// TIA Portal project "OP-TQ-01" (V13) (continued)
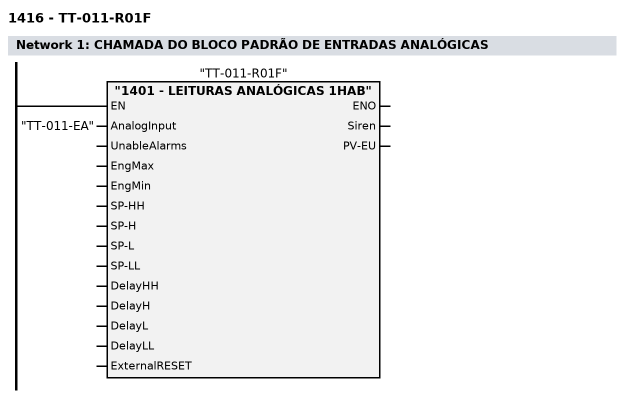
   RUNG wire#powerrail
      "TT-011-R01F"(AnalogInput := "TT-011-EA", UnableAlarms :=, EngMax :=, EngMin :=, "SP-HH" :=, "SP-H" :=, "SP-L" :=, "SP-LL" :=, DelayHH :=, DelayH :=, DelayL :=, DelayLL :=, ExternalRESET :=, Siren =>, "PV-EU" =>)
   END_RUNG
   // the same network as SCL:
   "TT-011-R01F"(AnalogInput := "TT-011-EA");   // "1401 - LEITURAS ANALÓGICAS 1HAB"
END_REGION
END_FUNCTION

// folder: PARAMETRIZADOS

FUNCTION_BLOCK "1110 - RESISTENCIAS"   // FB1110, LAD
{ S7_Optimized_Access := 'FALSE' }
VERSION : 0.1
   VAR_TEMP   // added for the SCL form of the ladder/FBD networks
      _w1 : Bool;
      _w2 : Bool;
   END_VAR
BEGIN

REGION Network 1: RESET FALHAS
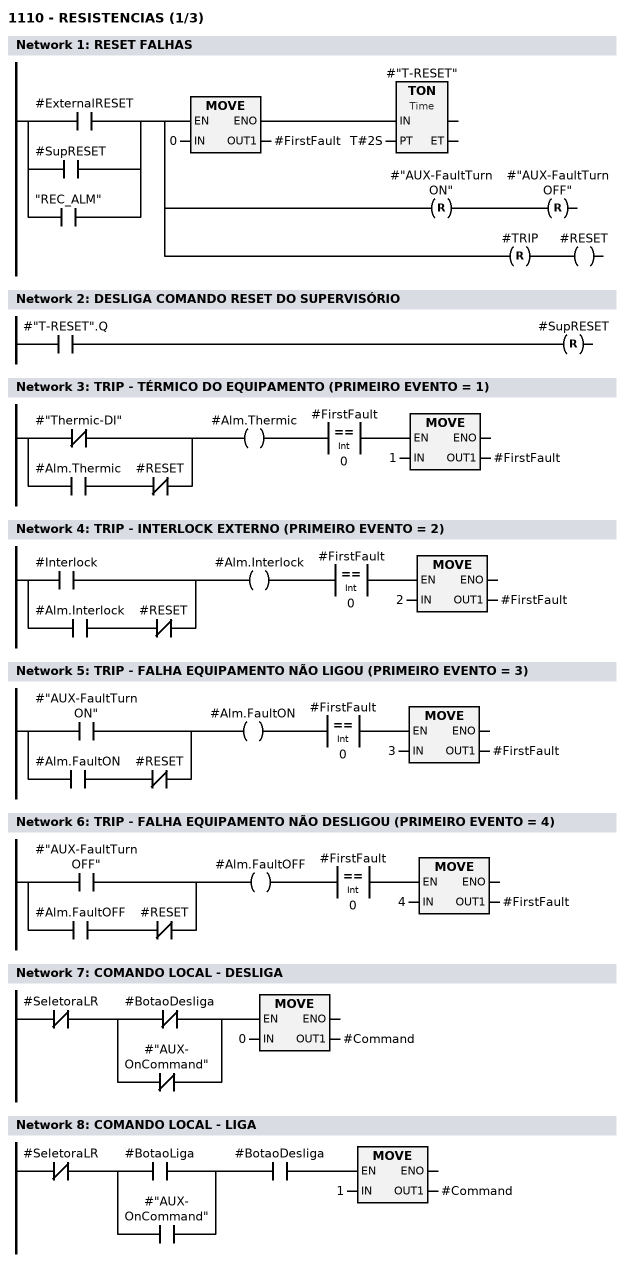
   // ENO of a box is taken as its EN; it also drops when the box reports an error
   #_w1 := #ExternalRESET OR #SupRESET OR "REC_ALM";
   IF #_w1 THEN #FirstFault := 0; END_IF;
   #"T-RESET".TON(IN := #_w1, PT := T#2S);
   IF #_w1 THEN
       #"AUX-FaultTurnON" := FALSE;
       #"AUX-FaultTurnOFF" := FALSE;
       #TRIP := FALSE;
   END_IF;
   #RESET := #_w1;
END_REGION

REGION Network 2: DESLIGA COMANDO RESET DO SUPERVISÓRIO
   RUNG wire#powerrail
      Contact( #"T-RESET".Q )
      R_Coil( #SupRESET )
   END_RUNG
   // the same network as SCL:
   IF #"T-RESET".Q THEN #SupRESET := FALSE; END_IF;
END_REGION

REGION Network 3: TRIP - TÉRMICO DO EQUIPAMENTO (PRIMEIRO EVENTO = 1)
   RUNG wire#powerrail
      I_Contact( #"Thermic-DI" )
      wire#w1
      Coil( #Alm.Thermic )
      { S7_Templates := "SrcType := Int" } EQ_Contact(in1 := #FirstFault, in2 := 0)
      { S7_GenerateENO := "TRUE" } Move(in := 1, out1 => #FirstFault)
   END_RUNG
   RUNG wire#powerrail
      Contact( #Alm.Thermic )
      I_Contact( #RESET )
   END_RUNG wire#w1
   // the same network as SCL:
   #Alm.Thermic := NOT #"Thermic-DI" OR (#Alm.Thermic AND NOT #RESET);
   IF #Alm.Thermic AND (#FirstFault = 0) THEN #FirstFault := 1; END_IF;
END_REGION

REGION Network 4: TRIP - INTERLOCK EXTERNO (PRIMEIRO EVENTO = 2)
   RUNG wire#powerrail
      Contact( #Interlock )
      wire#w1
      Coil( #Alm.Interlock )
      { S7_Templates := "SrcType := Int" } EQ_Contact(in1 := #FirstFault, in2 := 0)
      { S7_GenerateENO := "TRUE" } Move(in := 2, out1 => #FirstFault)
   END_RUNG
   RUNG wire#powerrail
      Contact( #Alm.Interlock )
      I_Contact( #RESET )
   END_RUNG wire#w1
   // the same network as SCL:
   #Alm.Interlock := #Interlock OR (#Alm.Interlock AND NOT #RESET);
   IF #Alm.Interlock AND (#FirstFault = 0) THEN #FirstFault := 2; END_IF;
END_REGION

REGION Network 5: TRIP - FALHA EQUIPAMENTO NÃO LIGOU (PRIMEIRO EVENTO = 3)
   RUNG wire#powerrail
      Contact( #"AUX-FaultTurnON" )
      wire#w1
      Coil( #Alm.FaultON )
      { S7_Templates := "SrcType := Int" } EQ_Contact(in1 := #FirstFault, in2 := 0)
      { S7_GenerateENO := "TRUE" } Move(in := 3, out1 => #FirstFault)
   END_RUNG
   RUNG wire#powerrail
      Contact( #Alm.FaultON )
      I_Contact( #RESET )
   END_RUNG wire#w1
   // the same network as SCL:
   #Alm.FaultON := #"AUX-FaultTurnON" OR (#Alm.FaultON AND NOT #RESET);
   IF #Alm.FaultON AND (#FirstFault = 0) THEN #FirstFault := 3; END_IF;
END_REGION

REGION Network 6: TRIP - FALHA EQUIPAMENTO NÃO DESLIGOU (PRIMEIRO EVENTO = 4)
   RUNG wire#powerrail
      Contact( #"AUX-FaultTurnOFF" )
      wire#w1
      Coil( #Alm.FaultOFF )
      { S7_Templates := "SrcType := Int" } EQ_Contact(in1 := #FirstFault, in2 := 0)
      { S7_GenerateENO := "TRUE" } Move(in := 4, out1 => #FirstFault)
   END_RUNG
   RUNG wire#powerrail
      Contact( #Alm.FaultOFF )
      I_Contact( #RESET )
   END_RUNG wire#w1
   // the same network as SCL:
   #Alm.FaultOFF := #"AUX-FaultTurnOFF" OR (#Alm.FaultOFF AND NOT #RESET);
   IF #Alm.FaultOFF AND (#FirstFault = 0) THEN #FirstFault := 4; END_IF;
END_REGION

REGION Network 7: COMANDO LOCAL - DESLIGA
   RUNG wire#powerrail
      I_Contact( #SeletoraLR )
      wire#w1
      I_Contact( #BotaoDesliga )
      wire#w2
      { S7_GenerateENO := "TRUE" } Move(in := 0, out1 => #Command)
   END_RUNG
   RUNG wire#w1
      I_Contact( #"AUX-OnCommand" )
   END_RUNG wire#w2
   // the same network as SCL:
   IF NOT #SeletoraLR AND (NOT #BotaoDesliga OR NOT #"AUX-OnCommand") THEN #Command := 0; END_IF;
END_REGION

REGION Network 8: COMANDO LOCAL - LIGA
   RUNG wire#powerrail
      I_Contact( #SeletoraLR )
      wire#w1
      Contact( #BotaoLiga )
      wire#w2
      Contact( #BotaoDesliga )
      { S7_GenerateENO := "TRUE" } Move(in := 1, out1 => #Command)
   END_RUNG
   RUNG wire#w1
      Contact( #"AUX-OnCommand" )
   END_RUNG wire#w2
   // the same network as SCL:
   IF NOT #SeletoraLR AND (#BotaoLiga OR #"AUX-OnCommand") AND #BotaoDesliga THEN #Command := 1; END_IF;
END_REGION

REGION Network 9: COMANDO LIGA EQUIPAMENTO
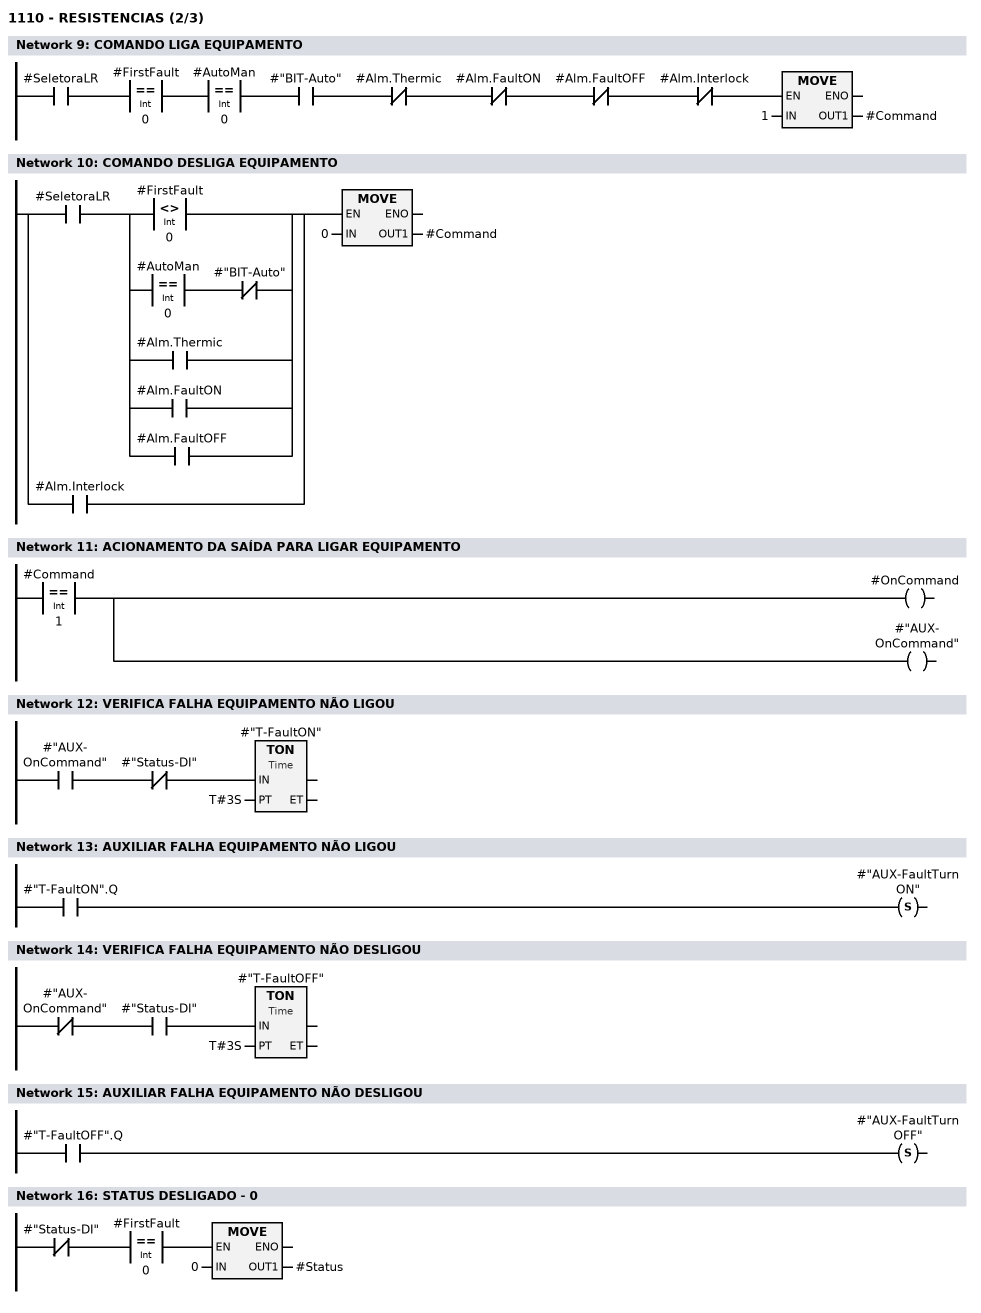
   RUNG wire#powerrail
      Contact( #SeletoraLR )
      { S7_Templates := "SrcType := Int" } EQ_Contact(in1 := #FirstFault, in2 := 0)
      { S7_Templates := "SrcType := Int" } EQ_Contact(in1 := #AutoMan, in2 := 0)
      Contact( #"BIT-Auto" )
      I_Contact( #Alm.Thermic )
      I_Contact( #Alm.FaultON )
      I_Contact( #Alm.FaultOFF )
      I_Contact( #Alm.Interlock )
      { S7_GenerateENO := "TRUE" } Move(in := 1, out1 => #Command)
   END_RUNG
   // the same network as SCL:
   IF #SeletoraLR AND (#FirstFault = 0) AND (#AutoMan = 0) AND #"BIT-Auto" AND NOT #Alm.Thermic AND NOT #Alm.FaultON AND NOT #Alm.FaultOFF AND NOT #Alm.Interlock THEN
       #Command := 1;
   END_IF;
END_REGION

REGION Network 10: COMANDO DESLIGA EQUIPAMENTO
   RUNG wire#powerrail
      Contact( #SeletoraLR )
      wire#w1
      { S7_Templates := "SrcType := Int" } NE_Contact(in1 := #FirstFault, in2 := 0)
      wire#w2
      { S7_GenerateENO := "TRUE" } Move(in := 0, out1 => #Command)
   END_RUNG
   RUNG wire#w1
      { S7_Templates := "SrcType := Int" } EQ_Contact(in1 := #AutoMan, in2 := 0)
      I_Contact( #"BIT-Auto" )
   END_RUNG wire#w2
   RUNG wire#w1
      Contact( #Alm.Thermic )
   END_RUNG wire#w2
   RUNG wire#w1
      Contact( #Alm.FaultON )
   END_RUNG wire#w2
   RUNG wire#w1
      Contact( #Alm.FaultOFF )
   END_RUNG wire#w2
   RUNG wire#powerrail
      Contact( #Alm.Interlock )
   END_RUNG wire#w2
   // the same network as SCL:
   IF (#SeletoraLR AND ((#FirstFault <> 0) OR ((#AutoMan = 0) AND NOT #"BIT-Auto") OR #Alm.Thermic OR #Alm.FaultON OR #Alm.FaultOFF)) OR #Alm.Interlock THEN
       #Command := 0;
   END_IF;
END_REGION

REGION Network 11: ACIONAMENTO DA SAÍDA PARA LIGAR EQUIPAMENTO
   RUNG wire#powerrail
      { S7_Templates := "SrcType := Int" } EQ_Contact(in1 := #Command, in2 := 1)
      wire#w1
      Coil( #OnCommand )
   END_RUNG
   RUNG wire#w1
      Coil( #"AUX-OnCommand" )
   END_RUNG
   // the same network as SCL:
   #OnCommand := #Command = 1;
   #"AUX-OnCommand" := #OnCommand;
END_REGION

REGION Network 12: VERIFICA FALHA EQUIPAMENTO NÃO LIGOU
   #"T-FaultON".TON(IN := #"AUX-OnCommand" AND NOT #"Status-DI", PT := T#3S);
END_REGION

REGION Network 13: AUXILIAR FALHA EQUIPAMENTO NÃO LIGOU
   RUNG wire#powerrail
      Contact( #"T-FaultON".Q )
      S_Coil( #"AUX-FaultTurnON" )
   END_RUNG
   // the same network as SCL:
   IF #"T-FaultON".Q THEN #"AUX-FaultTurnON" := TRUE; END_IF;
END_REGION

REGION Network 14: VERIFICA FALHA EQUIPAMENTO NÃO DESLIGOU
   #"T-FaultOFF".TON(IN := NOT #"AUX-OnCommand" AND #"Status-DI", PT := T#3S);
END_REGION

REGION Network 15: AUXILIAR FALHA EQUIPAMENTO NÃO DESLIGOU
   RUNG wire#powerrail
      Contact( #"T-FaultOFF".Q )
      S_Coil( #"AUX-FaultTurnOFF" )
   END_RUNG
   // the same network as SCL:
   IF #"T-FaultOFF".Q THEN #"AUX-FaultTurnOFF" := TRUE; END_IF;
END_REGION

REGION Network 16: STATUS DESLIGADO - 0
   RUNG wire#powerrail
      I_Contact( #"Status-DI" )
      { S7_Templates := "SrcType := Int" } EQ_Contact(in1 := #FirstFault, in2 := 0)
      { S7_GenerateENO := "TRUE" } Move(in := 0, out1 => #Status)
   END_RUNG
   // the same network as SCL:
   IF NOT #"Status-DI" AND (#FirstFault = 0) THEN #Status := 0; END_IF;
END_REGION

REGION Network 17: STATUS LIGADO - 1
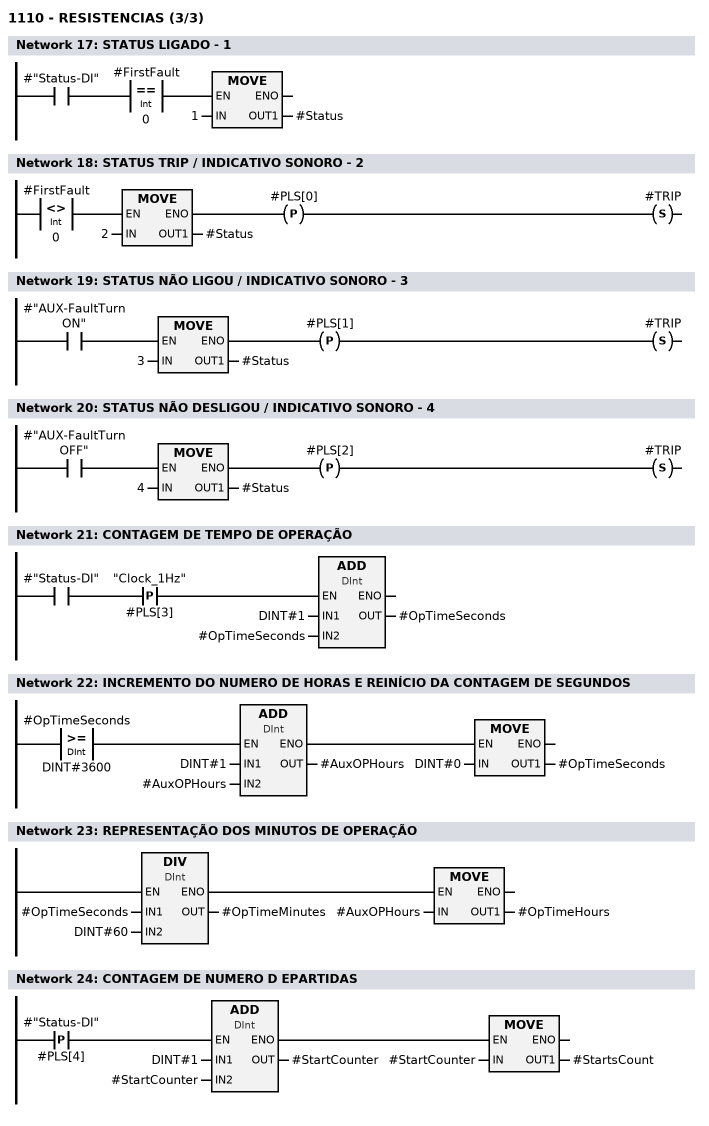
   RUNG wire#powerrail
      Contact( #"Status-DI" )
      { S7_Templates := "SrcType := Int" } EQ_Contact(in1 := #FirstFault, in2 := 0)
      { S7_GenerateENO := "TRUE" } Move(in := 1, out1 => #Status)
   END_RUNG
   // the same network as SCL:
   IF #"Status-DI" AND (#FirstFault = 0) THEN #Status := 1; END_IF;
END_REGION

REGION Network 18: STATUS TRIP / INDICATIVO SONORO - 2
   RUNG wire#powerrail
      { S7_Templates := "SrcType := Int" } NE_Contact(in1 := #FirstFault, in2 := 0)
      { S7_GenerateENO := "TRUE" } Move(in := 2, out1 => #Status)
      P_Trig( #PLS[0] )
      S_Coil( #TRIP )
   END_RUNG
   // the same network as SCL:
   // ENO of a box is taken as its EN; it also drops when the box reports an error
   #_w1 := #FirstFault <> 0;
   IF #_w1 THEN #Status := 2; END_IF;
   #_w2 := #_w1 AND NOT #PLS[0];   // rising edge
   #PLS[0] := #_w1;
   IF #_w2 THEN #TRIP := TRUE; END_IF;
END_REGION

REGION Network 19: STATUS NÃO LIGOU / INDICATIVO SONORO - 3
   RUNG wire#powerrail
      Contact( #"AUX-FaultTurnON" )
      { S7_GenerateENO := "TRUE" } Move(in := 3, out1 => #Status)
      P_Trig( #PLS[1] )
      S_Coil( #TRIP )
   END_RUNG
   // the same network as SCL:
   // ENO of a box is taken as its EN; it also drops when the box reports an error
   IF #"AUX-FaultTurnON" THEN #Status := 3; END_IF;
   #_w1 := #"AUX-FaultTurnON" AND NOT #PLS[1];   // rising edge
   #PLS[1] := #"AUX-FaultTurnON";
   IF #_w1 THEN #TRIP := TRUE; END_IF;
END_REGION

REGION Network 20: STATUS NÃO DESLIGOU / INDICATIVO SONORO - 4
   RUNG wire#powerrail
      Contact( #"AUX-FaultTurnOFF" )
      { S7_GenerateENO := "TRUE" } Move(in := 4, out1 => #Status)
      P_Trig( #PLS[2] )
      S_Coil( #TRIP )
   END_RUNG
   // the same network as SCL:
   // ENO of a box is taken as its EN; it also drops when the box reports an error
   IF #"AUX-FaultTurnOFF" THEN #Status := 4; END_IF;
   #_w1 := #"AUX-FaultTurnOFF" AND NOT #PLS[2];   // rising edge
   #PLS[2] := #"AUX-FaultTurnOFF";
   IF #_w1 THEN #TRIP := TRUE; END_IF;
END_REGION

REGION Network 21: CONTAGEM DE TEMPO DE OPERAÇÃO
   RUNG wire#powerrail
      Contact( #"Status-DI" )
      P_Contact(operand := "Clock_1Hz", bit := #PLS[3])
      { S7_Templates := "SrcType := DInt"; S7_GenerateENO := "TRUE" } Add(in1 := DINT#1, in2 := #OpTimeSeconds, out => #OpTimeSeconds)
   END_RUNG
   // the same network as SCL:
   #_w1 := #"Status-DI" AND "Clock_1Hz" AND NOT #PLS[3];   // rising edge of "Clock_1Hz"
   #PLS[3] := "Clock_1Hz";
   IF #_w1 THEN #OpTimeSeconds := DINT#1 + #OpTimeSeconds; END_IF;
END_REGION

REGION Network 22: INCREMENTO DO NUMERO DE HORAS E REINÍCIO DA CONTAGEM DE SEGUNDOS
   RUNG wire#powerrail
      { S7_Templates := "SrcType := DInt" } GE_Contact(in1 := #OpTimeSeconds, in2 := DINT#3600)
      { S7_Templates := "SrcType := DInt"; S7_GenerateENO := "TRUE" } Add(in1 := DINT#1, in2 := #AuxOPHours, out => #AuxOPHours)
      { S7_GenerateENO := "TRUE" } Move(in := DINT#0, out1 => #OpTimeSeconds)
   END_RUNG
   // the same network as SCL:
   // ENO of a box is taken as its EN; it also drops when the box reports an error
   IF #OpTimeSeconds >= DINT#3600 THEN
       #AuxOPHours := DINT#1 + #AuxOPHours;
       #OpTimeSeconds := DINT#0;
   END_IF;
END_REGION

REGION Network 23: REPRESENTAÇÃO DOS MINUTOS DE OPERAÇÃO
   RUNG wire#powerrail
      { S7_Templates := "SrcType := DInt"; S7_GenerateENO := "TRUE" } Div(in1 := #OpTimeSeconds, in2 := DINT#60, out => #OpTimeMinutes)
      { S7_GenerateENO := "TRUE" } Move(in := #AuxOPHours, out1 => #OpTimeHours)
   END_RUNG
   // the same network as SCL:
   // ENO of a box is taken as its EN; it also drops when the box reports an error
   #OpTimeMinutes := #OpTimeSeconds / DINT#60;
   #OpTimeHours := #AuxOPHours;
END_REGION

REGION Network 24: CONTAGEM DE NUMERO D EPARTIDAS
   RUNG wire#powerrail
      P_Contact(operand := #"Status-DI", bit := #PLS[4])
      { S7_Templates := "SrcType := DInt"; S7_GenerateENO := "TRUE" } Add(in1 := DINT#1, in2 := #StartCounter, out => #StartCounter)
      { S7_GenerateENO := "TRUE" } Move(in := #StartCounter, out1 => #StartsCount)
   END_RUNG
   // the same network as SCL:
   // ENO of a box is taken as its EN; it also drops when the box reports an error
   #_w1 := #"Status-DI" AND NOT #PLS[4];   // rising edge of #"Status-DI"
   #PLS[4] := #"Status-DI";
   IF #_w1 THEN
       #StartCounter := DINT#1 + #StartCounter;
       #StartsCount := #StartCounter;
   END_IF;
END_REGION
END_FUNCTION_BLOCK

FUNCTION_BLOCK "1401 - LEITURAS ANALÓGICAS 1HAB"   // FB1401, LAD
TITLE = LEITURA E VERIFICAÇÃO DE ALARMES ANALÓGICOS
{ S7_Optimized_Access := 'FALSE' }
VERSION : 0.1
   VAR_TEMP   // added for the SCL form of the ladder/FBD networks
      _w1 : Bool;
      _w2 : Bool;
      _w3 : Bool;
      _w4 : Bool;
   END_VAR
BEGIN

REGION Network 1: RESET FALHAS
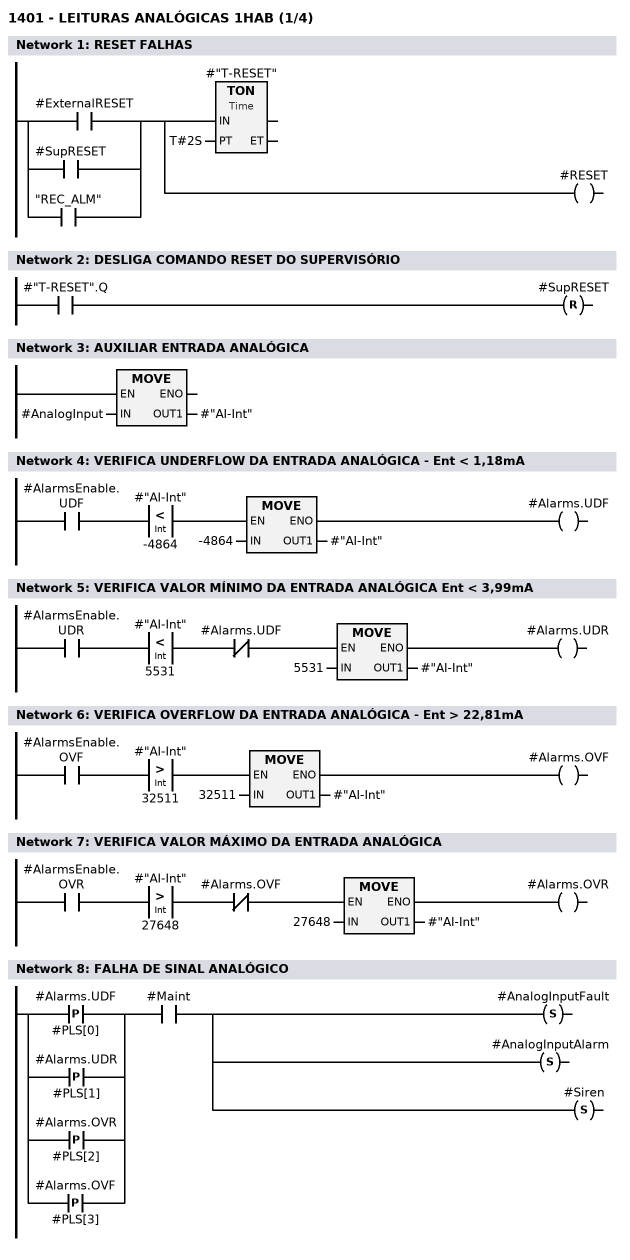
   #_w1 := #ExternalRESET OR #SupRESET OR "REC_ALM";
   #"T-RESET".TON(IN := #_w1, PT := T#2S);
   #RESET := #_w1;
END_REGION

REGION Network 2: DESLIGA COMANDO RESET DO SUPERVISÓRIO
   RUNG wire#powerrail
      Contact( #"T-RESET".Q )
      R_Coil( #SupRESET )
   END_RUNG
   // the same network as SCL:
   IF #"T-RESET".Q THEN #SupRESET := FALSE; END_IF;
END_REGION

REGION Network 3: AUXILIAR ENTRADA ANALÓGICA
   RUNG wire#powerrail
      { S7_GenerateENO := "TRUE" } Move(in := #AnalogInput, out1 => #"AI-Int")
   END_RUNG
   // the same network as SCL:
   #"AI-Int" := #AnalogInput;
END_REGION

REGION Network 4: VERIFICA UNDERFLOW DA ENTRADA ANALÓGICA - Ent < 1,18mA
   RUNG wire#powerrail
      Contact( #AlarmsEnable.UDF )
      { S7_Templates := "SrcType := Int" } LT_Contact(in1 := #"AI-Int", in2 := -4864)
      { S7_GenerateENO := "TRUE" } Move(in := -4864, out1 => #"AI-Int")
      Coil( #Alarms.UDF )
   END_RUNG
   // the same network as SCL:
   // ENO of a box is taken as its EN; it also drops when the box reports an error
   #_w1 := #AlarmsEnable.UDF AND (#"AI-Int" < (-4864));
   IF #_w1 THEN #"AI-Int" := -4864; END_IF;
   #Alarms.UDF := #_w1;
END_REGION

REGION Network 5: VERIFICA VALOR MÍNIMO DA ENTRADA ANALÓGICA Ent < 3,99mA
   RUNG wire#powerrail
      Contact( #AlarmsEnable.UDR )
      { S7_Templates := "SrcType := Int" } LT_Contact(in1 := #"AI-Int", in2 := 5531)
      I_Contact( #Alarms.UDF )
      { S7_GenerateENO := "TRUE" } Move(in := 5531, out1 => #"AI-Int")
      Coil( #Alarms.UDR )
   END_RUNG
   // the same network as SCL:
   // ENO of a box is taken as its EN; it also drops when the box reports an error
   #_w1 := #AlarmsEnable.UDR AND (#"AI-Int" < 5531) AND NOT #Alarms.UDF;
   IF #_w1 THEN #"AI-Int" := 5531; END_IF;
   #Alarms.UDR := #_w1;
END_REGION

REGION Network 6: VERIFICA OVERFLOW DA ENTRADA ANALÓGICA - Ent > 22,81mA
   RUNG wire#powerrail
      Contact( #AlarmsEnable.OVF )
      { S7_Templates := "SrcType := Int" } GT_Contact(in1 := #"AI-Int", in2 := 32511)
      { S7_GenerateENO := "TRUE" } Move(in := 32511, out1 => #"AI-Int")
      Coil( #Alarms.OVF )
   END_RUNG
   // the same network as SCL:
   // ENO of a box is taken as its EN; it also drops when the box reports an error
   #_w1 := #AlarmsEnable.OVF AND (#"AI-Int" > 32511);
   IF #_w1 THEN #"AI-Int" := 32511; END_IF;
   #Alarms.OVF := #_w1;
END_REGION

REGION Network 7: VERIFICA VALOR MÁXIMO DA ENTRADA ANALÓGICA
   RUNG wire#powerrail
      Contact( #AlarmsEnable.OVR )
      { S7_Templates := "SrcType := Int" } GT_Contact(in1 := #"AI-Int", in2 := 27648)
      I_Contact( #Alarms.OVF )
      { S7_GenerateENO := "TRUE" } Move(in := 27648, out1 => #"AI-Int")
      Coil( #Alarms.OVR )
   END_RUNG
   // the same network as SCL:
   // ENO of a box is taken as its EN; it also drops when the box reports an error
   #_w1 := #AlarmsEnable.OVR AND (#"AI-Int" > 27648) AND NOT #Alarms.OVF;
   IF #_w1 THEN #"AI-Int" := 27648; END_IF;
   #Alarms.OVR := #_w1;
END_REGION

REGION Network 8: FALHA DE SINAL ANALÓGICO
   RUNG wire#powerrail
      P_Contact(operand := #Alarms.UDF, bit := #PLS[0])
      wire#w1
      Contact( #Maint )
      wire#w2
      S_Coil( #AnalogInputFault )
   END_RUNG
   RUNG wire#powerrail
      P_Contact(operand := #Alarms.UDR, bit := #PLS[1])
   END_RUNG wire#w1
   RUNG wire#powerrail
      P_Contact(operand := #Alarms.OVR, bit := #PLS[2])
   END_RUNG wire#w1
   RUNG wire#powerrail
      P_Contact(operand := #Alarms.OVF, bit := #PLS[3])
   END_RUNG wire#w1
   RUNG wire#w2
      S_Coil( #AnalogInputAlarm )
   END_RUNG
   RUNG wire#w2
      S_Coil( #Siren )
   END_RUNG
   // the same network as SCL:
   #_w1 := #Alarms.UDF AND NOT #PLS[0];   // rising edge of #Alarms.UDF
   #PLS[0] := #Alarms.UDF;
   #_w2 := #Alarms.UDR AND NOT #PLS[1];   // rising edge of #Alarms.UDR
   #PLS[1] := #Alarms.UDR;
   #_w3 := #Alarms.OVR AND NOT #PLS[2];   // rising edge of #Alarms.OVR
   #PLS[2] := #Alarms.OVR;
   #_w4 := #Alarms.OVF AND NOT #PLS[3];   // rising edge of #Alarms.OVF
   #PLS[3] := #Alarms.OVF;
   IF (#_w1 OR #_w2 OR #_w3 OR #_w4) AND #Maint THEN
       #AnalogInputFault := TRUE;
       #AnalogInputAlarm := TRUE;
       #Siren := TRUE;
   END_IF;
END_REGION

REGION Network 9: RESET FALHA DE SINAL ANALÓGICO
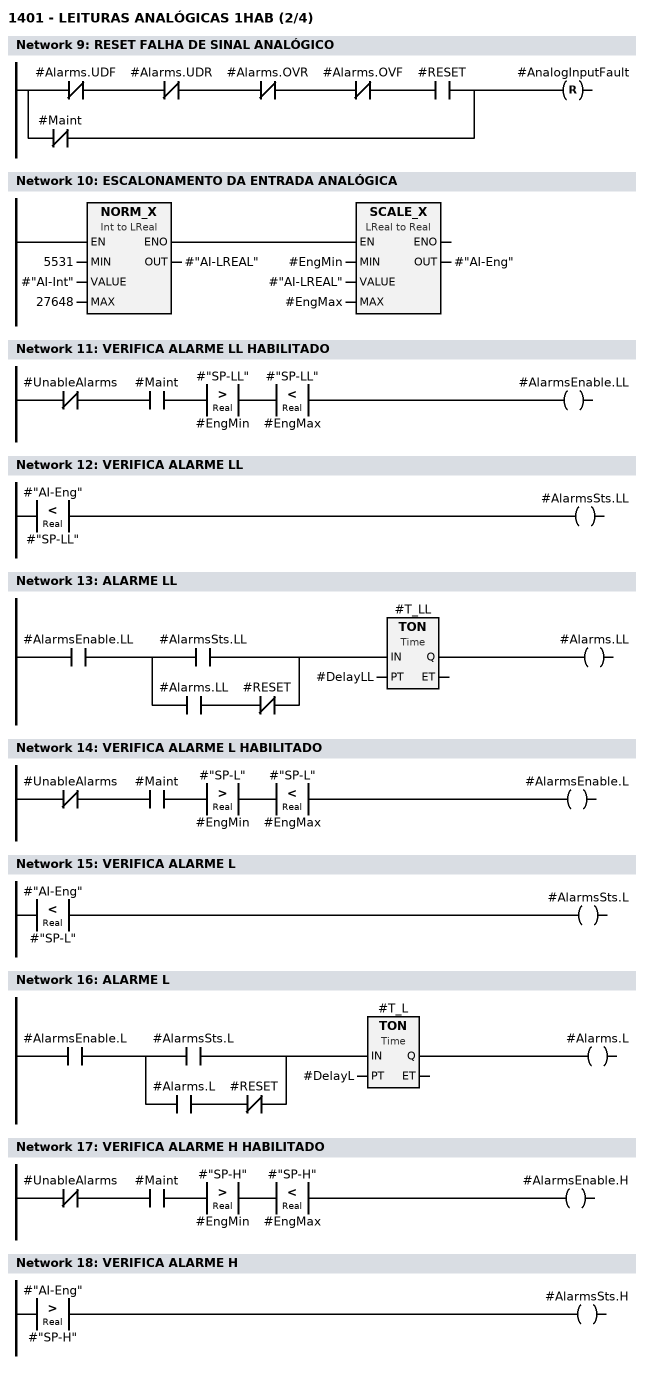
   RUNG wire#powerrail
      I_Contact( #Alarms.UDF )
      I_Contact( #Alarms.UDR )
      I_Contact( #Alarms.OVR )
      I_Contact( #Alarms.OVF )
      Contact( #RESET )
      wire#w1
      R_Coil( #AnalogInputFault )
   END_RUNG
   RUNG wire#powerrail
      I_Contact( #Maint )
   END_RUNG wire#w1
   // the same network as SCL:
   IF (NOT #Alarms.UDF AND NOT #Alarms.UDR AND NOT #Alarms.OVR AND NOT #Alarms.OVF AND #RESET) OR NOT #Maint THEN
       #AnalogInputFault := FALSE;
   END_IF;
END_REGION

REGION Network 10: ESCALONAMENTO DA ENTRADA ANALÓGICA
   RUNG wire#powerrail
      { S7_Templates := "[SrcType := Int, DestType := LReal]"; S7_GenerateENO := "TRUE" } Normalize(min := 5531, value := #"AI-Int", max := 27648, out => #"AI-LREAL")
      { S7_Templates := "[SrcType := LReal, DestType := Real]"; S7_GenerateENO := "TRUE" } Scale(min := #EngMin, value := #"AI-LREAL", max := #EngMax, out => #"AI-Eng")
   END_RUNG
   // the same network as SCL:
   // ENO of a box is taken as its EN; it also drops when the box reports an error
   #"AI-LREAL" := NORM_X(MIN := 5531, VALUE := #"AI-Int", MAX := 27648);
   #"AI-Eng" := SCALE_X(MIN := #EngMin, VALUE := #"AI-LREAL", MAX := #EngMax);
END_REGION

REGION Network 11: VERIFICA ALARME LL HABILITADO
   RUNG wire#powerrail
      I_Contact( #UnableAlarms )
      Contact( #Maint )
      { S7_Templates := "SrcType := Real" } GT_Contact(in1 := #"SP-LL", in2 := #EngMin)
      { S7_Templates := "SrcType := Real" } LT_Contact(in1 := #"SP-LL", in2 := #EngMax)
      Coil( #AlarmsEnable.LL )
   END_RUNG
   // the same network as SCL:
   #AlarmsEnable.LL := NOT #UnableAlarms AND #Maint AND (#"SP-LL" > #EngMin) AND (#"SP-LL" < #EngMax);
END_REGION

REGION Network 12: VERIFICA ALARME LL
   RUNG wire#powerrail
      { S7_Templates := "SrcType := Real" } LT_Contact(in1 := #"AI-Eng", in2 := #"SP-LL")
      Coil( #AlarmsSts.LL )
   END_RUNG
   // the same network as SCL:
   #AlarmsSts.LL := #"AI-Eng" < #"SP-LL";
END_REGION

REGION Network 13: ALARME LL
   #T_LL.TON(IN := #AlarmsEnable.LL AND (#AlarmsSts.LL OR (#Alarms.LL AND NOT #RESET)), PT := #DelayLL);
   #Alarms.LL := #T_LL.Q;
END_REGION

REGION Network 14: VERIFICA ALARME L HABILITADO
   RUNG wire#powerrail
      I_Contact( #UnableAlarms )
      Contact( #Maint )
      { S7_Templates := "SrcType := Real" } GT_Contact(in1 := #"SP-L", in2 := #EngMin)
      { S7_Templates := "SrcType := Real" } LT_Contact(in1 := #"SP-L", in2 := #EngMax)
      Coil( #AlarmsEnable.L )
   END_RUNG
   // the same network as SCL:
   #AlarmsEnable.L := NOT #UnableAlarms AND #Maint AND (#"SP-L" > #EngMin) AND (#"SP-L" < #EngMax);
END_REGION

REGION Network 15: VERIFICA ALARME L
   RUNG wire#powerrail
      { S7_Templates := "SrcType := Real" } LT_Contact(in1 := #"AI-Eng", in2 := #"SP-L")
      Coil( #AlarmsSts.L )
   END_RUNG
   // the same network as SCL:
   #AlarmsSts.L := #"AI-Eng" < #"SP-L";
END_REGION

REGION Network 16: ALARME L
   #T_L.TON(IN := #AlarmsEnable.L AND (#AlarmsSts.L OR (#Alarms.L AND NOT #RESET)), PT := #DelayL);
   #Alarms.L := #T_L.Q;
END_REGION

REGION Network 17: VERIFICA ALARME H HABILITADO
   RUNG wire#powerrail
      I_Contact( #UnableAlarms )
      Contact( #Maint )
      { S7_Templates := "SrcType := Real" } GT_Contact(in1 := #"SP-H", in2 := #EngMin)
      { S7_Templates := "SrcType := Real" } LT_Contact(in1 := #"SP-H", in2 := #EngMax)
      Coil( #AlarmsEnable.H )
   END_RUNG
   // the same network as SCL:
   #AlarmsEnable.H := NOT #UnableAlarms AND #Maint AND (#"SP-H" > #EngMin) AND (#"SP-H" < #EngMax);
END_REGION

REGION Network 18: VERIFICA ALARME H
   RUNG wire#powerrail
      { S7_Templates := "SrcType := Real" } GT_Contact(in1 := #"AI-Eng", in2 := #"SP-H")
      Coil( #AlarmsSts.H )
   END_RUNG
   // the same network as SCL:
   #AlarmsSts.H := #"AI-Eng" > #"SP-H";
END_REGION

REGION Network 19: ALARME H
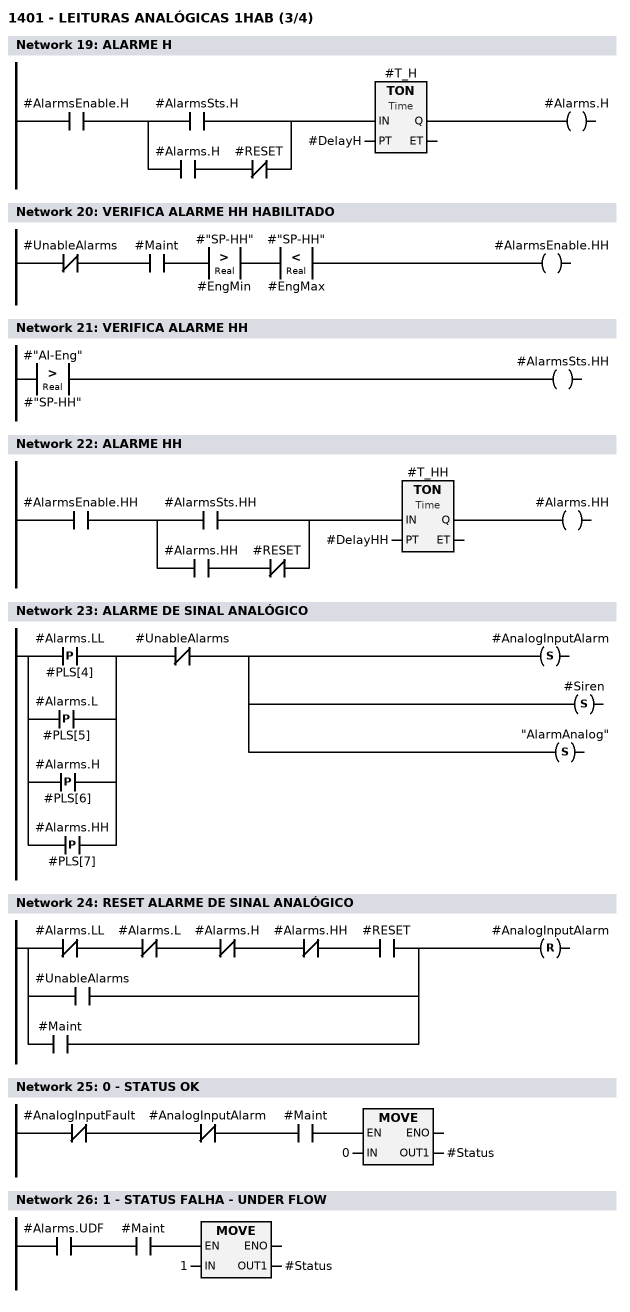
   #T_H.TON(IN := #AlarmsEnable.H AND (#AlarmsSts.H OR (#Alarms.H AND NOT #RESET)), PT := #DelayH);
   #Alarms.H := #T_H.Q;
END_REGION

REGION Network 20: VERIFICA ALARME HH HABILITADO
   RUNG wire#powerrail
      I_Contact( #UnableAlarms )
      Contact( #Maint )
      { S7_Templates := "SrcType := Real" } GT_Contact(in1 := #"SP-HH", in2 := #EngMin)
      { S7_Templates := "SrcType := Real" } LT_Contact(in1 := #"SP-HH", in2 := #EngMax)
      Coil( #AlarmsEnable.HH )
   END_RUNG
   // the same network as SCL:
   #AlarmsEnable.HH := NOT #UnableAlarms AND #Maint AND (#"SP-HH" > #EngMin) AND (#"SP-HH" < #EngMax);
END_REGION

REGION Network 21: VERIFICA ALARME HH
   RUNG wire#powerrail
      { S7_Templates := "SrcType := Real" } GT_Contact(in1 := #"AI-Eng", in2 := #"SP-HH")
      Coil( #AlarmsSts.HH )
   END_RUNG
   // the same network as SCL:
   #AlarmsSts.HH := #"AI-Eng" > #"SP-HH";
END_REGION

REGION Network 22: ALARME HH
   #T_HH.TON(IN := #AlarmsEnable.HH AND (#AlarmsSts.HH OR (#Alarms.HH AND NOT #RESET)), PT := #DelayHH);
   #Alarms.HH := #T_HH.Q;
END_REGION

REGION Network 23: ALARME DE SINAL ANALÓGICO
   RUNG wire#powerrail
      P_Contact(operand := #Alarms.LL, bit := #PLS[4])
      wire#w1
      I_Contact( #UnableAlarms )
      wire#w2
      S_Coil( #AnalogInputAlarm )
   END_RUNG
   RUNG wire#powerrail
      P_Contact(operand := #Alarms.L, bit := #PLS[5])
   END_RUNG wire#w1
   RUNG wire#powerrail
      P_Contact(operand := #Alarms.H, bit := #PLS[6])
   END_RUNG wire#w1
   RUNG wire#powerrail
      P_Contact(operand := #Alarms.HH, bit := #PLS[7])
   END_RUNG wire#w1
   RUNG wire#w2
      S_Coil( #Siren )
   END_RUNG
   RUNG wire#w2
      S_Coil( "AlarmAnalog" )
   END_RUNG
   // the same network as SCL:
   #_w1 := #Alarms.LL AND NOT #PLS[4];   // rising edge of #Alarms.LL
   #PLS[4] := #Alarms.LL;
   #_w2 := #Alarms.L AND NOT #PLS[5];   // rising edge of #Alarms.L
   #PLS[5] := #Alarms.L;
   #_w3 := #Alarms.H AND NOT #PLS[6];   // rising edge of #Alarms.H
   #PLS[6] := #Alarms.H;
   #_w4 := #Alarms.HH AND NOT #PLS[7];   // rising edge of #Alarms.HH
   #PLS[7] := #Alarms.HH;
   IF (#_w1 OR #_w2 OR #_w3 OR #_w4) AND NOT #UnableAlarms THEN
       #AnalogInputAlarm := TRUE;
       #Siren := TRUE;
       "AlarmAnalog" := TRUE;
   END_IF;
END_REGION
